// TIA Portal project "Vent_Fan_PLC_202203231" (V16)

(* hardware
DEVICE "ET 200SP station_1"  ET 200SP-Station
   slot 0: "Rack_0"  Rack  6ES5 710-8MAx1
   slot 1: "Roof Fans PLC"  CPU 1512SP-1 PN  6ES7 512-1DK01-0AB0  V2.1
      slot 32768: "PROFINET interface_1"  X1
         slot 32771: "Port_3"  X1 P3
   slot 2: "DI 16x24VDC ST_1"  DI 16x24VDC ST  6ES7 131-6BH00-0BA0  V1.1
      slot 1: "DI 16x24VDC ST_1"  DI 16x24VDC ST
   slot 3: "DQ 16x24VDC/0.5A ST_1"  DQ 16x24VDC/0.5A ST  6ES7 132-6BH00-0BA0  V1.0
      slot 1: "DQ 16x24VDC/0.5A ST_1"  DQ 16x24VDC/0.5A ST
   slot 4: "Server module_1"  Server module  6ES7 193-6PA00-0AA0  V1.1
      slot 1: "Server module_1"  Server module
   slot 127: "BA 2xRJ45"  BA 2xRJ45  6ES7 193-6AR00-0AA0  V0.0
      slot 32769: "Port_1"  X1 P1  6ES7 193-6AR00-0AA0
      slot 32770: "Port_2"  X1 P2  6ES7 193-6AR00-0AA0
DEVICE "SINAMICS G_1"  Sinamics.Device
   slot 0: "	_0"  Rail  SinamicsG120CRackP
   slot 0: "RTU-0035"  G120C PN  6SL3210-1KE15-8UF2  4.7.10
      slot 1: "PROFINET interface"  MDD-SinamicsG120-P
      slot 3: "PM G120C"  PM G120C  6SL3210-1KE15-8UF2  -
DEVICE "SINAMICS G_2"  Sinamics.Device
   slot 0: "	_0"  Rail  SinamicsG120CRackP
   slot 0: "RTU-0010"  G120C PN  6SL3210-1KE15-8UF2  4.7.10
      slot 1: "PROFINET interface"  MDD-SinamicsG120-P
      slot 3: "PM G120C"  PM G120C  6SL3210-1KE15-8UF2  -
DEVICE "SINAMICS G_3"  Sinamics.Device
   slot 0: "	_0"  Rail  SinamicsG120CRackP
   slot 0: "RTU-0011"  G120C PN  6SL3210-1KE15-8UF2  4.7.10
      slot 1: "PROFINET interface"  MDD-SinamicsG120-P
      slot 3: "PM G120C"  PM G120C  6SL3210-1KE15-8UF2  -
DEVICE "SINAMICS G_4"  Sinamics.Device
   slot 0: "	_0"  Rail  SinamicsG120CRackP
   slot 0: "RTU-0014"  G120C PN  6SL3210-1KE15-8UF2  4.7.10
      slot 1: "PROFINET interface"  MDD-SinamicsG120-P
      slot 3: "PM G120C"  PM G120C  6SL3210-1KE15-8UF2  -
DEVICE "SINAMICS G_5"  Sinamics.Device
   slot 0: "	_0"  Rail  SinamicsG120CRackP
   slot 0: "RTU-0015"  G120C PN  6SL3210-1KE15-8UF2  4.7.10
      slot 1: "PROFINET interface"  MDD-SinamicsG120-P
      slot 3: "PM G120C"  PM G120C  6SL3210-1KE15-8UF2  -
DEVICE "SINAMICS G_6"  Sinamics.Device
   slot 0: "	_0"  Rail  SinamicsG120CRackP
   slot 0: "RTU-0020"  G120C PN  6SL3210-1KE15-8UF2  4.7.10
      slot 1: "PROFINET interface"  MDD-SinamicsG120-P
      slot 3: "PM G120C"  PM G120C  6SL3210-1KE15-8UF2  -
DEVICE "SINAMICS G_7"  Sinamics.Device
   slot 0: "	_0"  Rail  SinamicsG120CRackP
   slot 0: "RTU-0021"  G120C PN  6SL3210-1KE15-8UF2  4.7.10
      slot 1: "PROFINET interface"  MDD-SinamicsG120-P
      slot 3: "PM G120C"  PM G120C  6SL3210-1KE15-8UF2  -
DEVICE "SINAMICS G_8"  Sinamics.Device
   slot 0: "	_0"  Rail  SinamicsG120CRackP
   slot 0: "RTU-0052"  G120C PN  6SL3210-1KE15-8UF2  4.7.10
      slot 1: "PROFINET interface"  MDD-SinamicsG120-P
      slot 3: "PM G120C"  PM G120C  6SL3210-1KE15-8UF2  -
DEVICE "SINAMICS G_9"  Sinamics.Device
   slot 0: "	_0"  Rail  SinamicsG120CRackP
   slot 0: "RTU-0053"  G120C PN  6SL3210-1KE15-8UF2  4.7.10
      slot 1: "PROFINET interface"  MDD-SinamicsG120-P
      slot 3: "PM G120C"  PM G120C  6SL3210-1KE15-8UF2  -
DEVICE "SINAMICS G_10"  Sinamics.Device
   slot 0: "	_0"  Rail  SinamicsG120CRackP
   slot 0: "RTU-0054"  G120C PN  6SL3210-1KE15-8UF2  4.7.10
      slot 1: "PROFINET interface"  MDD-SinamicsG120-P
      slot 3: "PM G120C"  PM G120C  6SL3210-1KE15-8UF2  -
DEVICE "SINAMICS G_11"  Sinamics.Device
   slot 0: "	_0"  Rail  SinamicsG120CRackP
   slot 0: "RTU-0055"  G120C PN  6SL3210-1KE15-8UF2  4.7.10
      slot 1: "PROFINET interface"  MDD-SinamicsG120-P
      slot 3: "PM G120C"  PM G120C  6SL3210-1KE15-8UF2  -
DEVICE "SINAMICS G_12"  Sinamics.Device
   slot 0: "	_0"  Rail  SinamicsG120CRackP
   slot 0: "RTU-0042"  G120C PN  6SL3210-1KE15-8UF2  4.7.10
      slot 1: "PROFINET interface"  MDD-SinamicsG120-P
      slot 3: "PM G120C"  PM G120C  6SL3210-1KE15-8UF2  -
*)

// ===== PLC "Roof Fans PLC"  CPU 1512SP-1 PN =====

VAR_GLOBAL   // PLC tag table "Default tag table"
   "System_Byte" AT %MB1 : Byte;
   "FirstScan" AT %M1.0 : Bool;
   "DiagStatusUpdate" AT %M1.1 : Bool;
   "AlwaysTRUE" AT %M1.2 : Bool;
   "AlwaysFALSE" AT %M1.3 : Bool;
   "Clock_Byte" AT %MB0 : Byte;
   "Clock_10Hz" AT %M0.0 : Bool;
   "Clock_5Hz" AT %M0.1 : Bool;
   "Clock_2.5Hz" AT %M0.2 : Bool;
   "Clock_2Hz" AT %M0.3 : Bool;
   "Clock_1.25Hz" AT %M0.4 : Bool;
   "Clock_1Hz" AT %M0.5 : Bool;
   "Clock_0.625Hz" AT %M0.6 : Bool;
   "Clock_0.5Hz" AT %M0.7 : Bool;
   "Drive_Temp" AT %MD100 : Real;
END_VAR

VAR_GLOBAL CONSTANT   // PLC tag table "Default tag table"
   "STATION_COUNT" : Int := 49;   // 0 indexed
   "SCHEDULES_PER_DAY" : Int := 4;   // 0 indexed
   "TIME_STRING_LENGTH" : Int := 20;   // standard indexed
END_VAR

VAR_GLOBAL   // PLC tag table "INPUTS"
   "Input_1" AT %I0.0 : Bool;
   "Input_2" AT %I0.2 : Bool;
   "Input_3" AT %I0.3 : Bool;
   "Input_4" AT %I0.4 : Bool;
   "Input_5" AT %I0.5 : Bool;
   "Input_6" AT %I0.6 : Bool;
   "Input_7" AT %I0.7 : Bool;
   "Input_8" AT %I1.0 : Bool;
   "Input_9" AT %I1.1 : Bool;
   "Input_10" AT %I1.2 : Bool;
   "Input_11" AT %I1.3 : Bool;
   "Input_12" AT %I1.4 : Bool;
   "Input_13" AT %I1.5 : Bool;
   "Input_14" AT %I1.6 : Bool;
   "Input_15" AT %I1.7 : Bool;
END_VAR

VAR_GLOBAL   // PLC tag table "OUTPUTS"
   "Output_1" AT %Q0.0 : Bool;
   "Output_15" AT %Q1.6 : Bool;
   "Output_2" AT %Q0.1 : Bool;
   "Output_3" AT %Q0.2 : Bool;
   "Output_4" AT %Q0.3 : Bool;
   "Output_5" AT %Q0.4 : Bool;
   "Output_6" AT %Q0.5 : Bool;
   "Output_7" AT %Q0.6 : Bool;
   "Output_8" AT %Q0.7 : Bool;
   "Output_9" AT %Q1.0 : Bool;
   "Output_10" AT %Q1.1 : Bool;
   "Output_11" AT %Q1.2 : Bool;
   "Output_12" AT %Q1.3 : Bool;
   "Output_13" AT %Q1.4 : Bool;
   "Output_14" AT %Q1.5 : Bool;
END_VAR

VAR_GLOBAL   // PLC tag table "RTU-0035"
   "RTU-0035_Temperature" AT %IW260 : Word;
   "RTU-0035_Speed" AT %IW258 : Word;
   "RTU-0035_Current" AT %IW262 : Word;
END_VAR

VAR_GLOBAL   // PLC tag table "RTU-0010"
   "RTU-0010_Temperature" AT %IW268 : Word;
   "RTU-0010_Speed" AT %IW266 : Word;
   "RTU-0010_Current" AT %IW270 : Word;
END_VAR

VAR_GLOBAL   // PLC tag table "RTU-0011"
   "RTU-0011_Temperature" AT %IW276 : Word;
   "RTU-0011_Speed" AT %IW274 : Word;
   "RTU-0011_Current" AT %IW278 : Word;
END_VAR

VAR_GLOBAL   // PLC tag table "RTU-0014"
   "RTU-0014_Temperature" AT %IW284 : Word;
   "RTU-0014_Speed" AT %IW282 : Word;
   "RTU-0014_Current" AT %IW286 : Word;
END_VAR

VAR_GLOBAL   // PLC tag table "RTU-0015"
   "RTU-0015_Temperature" AT %IW292 : Word;
   "RTU-0015_Speed" AT %IW290 : Word;
   "RTU-0015_Current" AT %IW294 : Word;
END_VAR

VAR_GLOBAL   // PLC tag table "RTU-0020"
   "RTU-0020_Temperature" AT %IW300 : Word;
   "RTU-0020_Speed" AT %IW298 : Word;
   "RTU-0020_Current" AT %IW302 : Word;
END_VAR

VAR_GLOBAL   // PLC tag table "RTU-0021"
   "RTU-0021_Temperature" AT %IW308 : Word;
   "RTU-0021_Speed" AT %IW2306 : Word;
   "RTU-0021_Current" AT %IW310 : Word;
END_VAR

VAR_GLOBAL   // PLC tag table "RTU-0052"
   "RTU-0052_Temperature" AT %IW316 : Word;
   "RTU-0052_Speed" AT %IW314 : Word;
   "RTU-0052_Current" AT %IW318 : Word;
END_VAR

VAR_GLOBAL   // PLC tag table "RTU-0053"
   "RTU-0053_Temperature" AT %IW324 : Word;
   "RTU-0053_Speed" AT %IW322 : Word;
   "RTU-0053_Current" AT %IW326 : Word;
END_VAR

VAR_GLOBAL   // PLC tag table "RTU-0054"
   "RTU-0054_Temperature" AT %IW332 : Word;
   "RTU-0054_Speed" AT %IW330 : Word;
   "RTU-0054_Current" AT %IW334 : Word;
END_VAR

VAR_GLOBAL   // PLC tag table "RTU-0055"
   "RTU-0055_Temperature" AT %IW340 : Word;
   "RTU-0055_Speed" AT %IW338 : Word;
   "RTU-0055_Current" AT %IW342 : Word;
END_VAR

VAR_GLOBAL   // PLC tag table "RTU-0042"
   "RTU-0042_Temperature" AT %IW348 : Word;
   "RTU-0042_Speed" AT %IW346 : Word;
   "RTU-0042_Current" AT %IW350 : Word;
END_VAR

TYPE "Web_Meta.UDT"
   STRUCT
      drive : "Drive.UDT";
      faults : "Faults.UDT";
      id : Int;
      manual : "Station.Web_Interface.Manual.UDT";
      selected_station : Int;
      scheduled_speed : Real;
      temporal_schedule : "Web_Meta.Web_Interface.Schedules.Temporal.UDT";
      thermal_schedule : "Schedules.Thermal.UDT";
   END_STRUCT;
END_TYPE

TYPE "Sensors.Thermal.UDT"
   STRUCT
      me : "Convert.Word_to_Real.UDT";
   END_STRUCT;
END_TYPE

TYPE "Sensors.UDT"
   STRUCT
      thermal : "Sensors.Thermal.UDT";
   END_STRUCT;
END_TYPE

TYPE "Drive.UDT"
   STRUCT
      commands : "Drive.Commands.UDT";
      commands_manual : "Drive.Commands.UDT";
      commands_thermal : "Drive.Commands.UDT";
      commands_temporal : "Drive.Commands.UDT";
      feedback : "Drive.Feedback.UDT";
      sensors : "Sensors.UDT";
   END_STRUCT;
END_TYPE

TYPE "Stations.UDT"
   STRUCT
      me : Array[0.."STATION_COUNT"] of "Station.UDT";
   END_STRUCT;
   // me[7].drive.sensors.thermal.me.processed := 76.8;
   // me[7].drive.feedback.speed.me.processed := 1100.56;
   // me[7].drive.feedback.current.me.processed := 3.78;
END_TYPE

TYPE "Station.UDT"
   STRUCT
      drive : "Drive.UDT";
      faults : "Faults.UDT";
      interface : "Interface.UDT";
      schedules : "Schedules.UDT";
   END_STRUCT;
END_TYPE

TYPE "Drive.Feedback.UDT"
   STRUCT
      faults : String := 'none';
      current : "Drive.Feedback.Current.UDT";
      speed : "Drive.Feedback.Speed.UDT";
      state : String := 'not running';
   END_STRUCT;
END_TYPE

TYPE "Convert.Word_to_Real.UDT"
   STRUCT
      raw : Word;
      processed : Real;
   END_STRUCT;
END_TYPE

TYPE "Drive.Feedback.Speed.UDT"
   STRUCT
      me : "Convert.Word_to_Real.UDT";
   END_STRUCT;
END_TYPE

TYPE "Drive.Feedback.Current.UDT"
   STRUCT
      me : "Convert.Word_to_Real.UDT";
   END_STRUCT;
END_TYPE

TYPE "Station.Web_Interface.UDT"
   STRUCT
      manual : "Station.Web_Interface.Manual.UDT";
      temporal : "Web_Meta.Web_Interface.Schedules.Temporal.UDT";
   END_STRUCT;
END_TYPE

TYPE "Station.Web_Interface.Manual.UDT"
   STRUCT
      acknowledge : Bool;
      command_speed : Real;
      mode : String[20] := 'stop';
      override : Bool;
      submit : Bool;
      toggle : Bool;
   END_STRUCT;
END_TYPE

TYPE "Schedules.Thermal.Element.UDT"
   STRUCT
      temperature : Real;
      speed : Real;
   END_STRUCT;
END_TYPE

TYPE "Schedules.Thermal.UDT"
   STRUCT
      start : "Schedules.Thermal.Element.UDT";
      max : "Schedules.Thermal.Element.UDT";
   END_STRUCT;
END_TYPE

TYPE "Schedules.UDT"
   STRUCT
      thermal : "Schedules.Thermal.UDT";
      temporal : "Schedules.Temporal.UDT";
   END_STRUCT;
END_TYPE

TYPE "Web_Meta.Web_Interface.Schedules.Temporal.Element.UDT"
   STRUCT
      start : String["TIME_STRING_LENGTH"];
      stop : String["TIME_STRING_LENGTH"];
      speed : Real;
   END_STRUCT;
END_TYPE

TYPE "Faults.UDT"
   STRUCT
      color : String[6];
      fault : String;
   END_STRUCT;
END_TYPE

TYPE "Interface.UDT"
   STRUCT
      current_feedback_b0 : DInt;
      id : USInt;
      raw_temp_sensor_b0 : DInt;
      sensor_max_temp : Real := 150.0;
      sensor_min_temp : Real;
      speed_feedback_b0 : DInt;
      max_speed : Real := 1500.0;
      profinet_pointer_to_drive : Hw_SubModule;
   END_STRUCT;
END_TYPE

TYPE "Interface.Thermal.UDT"
   STRUCT
      pointer_to_raw_value : DInt;   // input word number of data from drive
      min : Real;
      max : Real := 150.0;
   END_STRUCT;
END_TYPE

TYPE "Interface.Drive.Feedback.UDT"
   STRUCT
      current : DInt;   // pointer to input word with raw value
      speed : DInt;   // pointer to input word with raw value
   END_STRUCT;
END_TYPE

TYPE "Interface.Sensors.UDT"
   STRUCT
      thermal : "Interface.Thermal.UDT";
   END_STRUCT;
END_TYPE

TYPE "Drive.Commands.UDT"
   STRUCT
      override : Bool;
      run : Bool;
      speed : Real;
      stop : Bool;
   END_STRUCT;
END_TYPE

TYPE "Interface.Drive.Settings.UTD"
   STRUCT
      id : Bool;
      profinet_pointer_to_drive : Hw_SubModule;
      max_speed : Real := 1500.0;
   END_STRUCT;
END_TYPE

TYPE "OPC.Station.UDT"
   STRUCT
      current : Real;
      id : USInt;
      speed : Real;
      temperature : Real;
   END_STRUCT;
END_TYPE

TYPE "OPC.Stations.UDT"
   STRUCT
      me : Array[0.."STATION_COUNT"] of "OPC.Station.UDT";
   END_STRUCT;
END_TYPE

TYPE "Web_Meta.Web_Interface.Schedules.Temporal.UDT"
   STRUCT
      monday : Array[0.."SCHEDULES_PER_DAY"] of "Web_Meta.Web_Interface.Schedules.Temporal.Element.UDT";
      tuesday : Array[0.."SCHEDULES_PER_DAY"] of "Web_Meta.Web_Interface.Schedules.Temporal.Element.UDT";
      wednesday : Array[0.."SCHEDULES_PER_DAY"] of "Web_Meta.Web_Interface.Schedules.Temporal.Element.UDT";
      thursday : Array[0.."SCHEDULES_PER_DAY"] of "Web_Meta.Web_Interface.Schedules.Temporal.Element.UDT";
      friday : Array[0.."SCHEDULES_PER_DAY"] of "Web_Meta.Web_Interface.Schedules.Temporal.Element.UDT";
      saturday : Array[0.."SCHEDULES_PER_DAY"] of "Web_Meta.Web_Interface.Schedules.Temporal.Element.UDT";
      sunday : Array[0.."SCHEDULES_PER_DAY"] of "Web_Meta.Web_Interface.Schedules.Temporal.Element.UDT";
      new_data : Bool;
   END_STRUCT;
END_TYPE

TYPE "Schedules.Temporal.UDT"
   STRUCT
      monday : Array[0.."SCHEDULES_PER_DAY"] of "Schedules.Temporal.Element.UDT";
      tuesday : Array[0.."SCHEDULES_PER_DAY"] of "Schedules.Temporal.Element.UDT";
      wednesday : Array[0.."SCHEDULES_PER_DAY"] of "Schedules.Temporal.Element.UDT";
      thursday : Array[0.."SCHEDULES_PER_DAY"] of "Schedules.Temporal.Element.UDT";
      friday : Array[0.."SCHEDULES_PER_DAY"] of "Schedules.Temporal.Element.UDT";
      saturday : Array[0.."SCHEDULES_PER_DAY"] of "Schedules.Temporal.Element.UDT";
      sunday : Array[0.."SCHEDULES_PER_DAY"] of "Schedules.Temporal.Element.UDT";
   END_STRUCT;
END_TYPE

TYPE "Schedules.Temporal.Element.Date_Time.UDT"
   STRUCT
      month : USInt;
      day : USInt;
      weekday : USInt;
      hour : USInt;
      minute : USInt;
   END_STRUCT;
END_TYPE

TYPE "Schedules.Temporal.Element.UDT"
   STRUCT
      start : "Schedules.Temporal.Element.Date_Time.UDT";
      stop : "Schedules.Temporal.Element.Date_Time.UDT";
      speed : Real;
   END_STRUCT;
END_TYPE

DATA_BLOCK "Web_Meta"   // DB1
{ S7_Optimized_Access := 'TRUE' }
VERSION : 0.1
BEGIN
END_DATA_BLOCK

DATA_BLOCK "Stations"   // DB2
{ S7_Optimized_Access := 'TRUE' }
VERSION : 0.1
BEGIN
   me[7].interface.id := 42;
   me[0].interface.id := 10;
   me[1].interface.id := 11;
   me[2].interface.id := 14;
   me[8].interface.id := 52;
   me[3].interface.id := 15;
   me[5].interface.id := 21;
   me[6].interface.id := 35;
   me[4].interface.id := 20;
   me[9].interface.id := 53;
   me[10].interface.id := 54;
   me[11].interface.id := 55;
   me[6].interface.current_feedback_b0 := 262;
   me[6].interface.raw_temp_sensor_b0 := 260;
   me[6].interface.sensor_max_temp := 150.0;
   me[6].interface.speed_feedback_b0 := 258;
   me[6].interface.max_speed := 1500.0;
   me[6].interface.profinet_pointer_to_drive := 269;
   me[0].interface.current_feedback_b0 := 270;
   me[0].interface.raw_temp_sensor_b0 := 268;
   me[0].interface.speed_feedback_b0 := 266;
   me[0].interface.profinet_pointer_to_drive := 278;
   me[1].interface.profinet_pointer_to_drive := 287;
   me[1].interface.speed_feedback_b0 := 274;
   me[1].interface.raw_temp_sensor_b0 := 276;
   me[1].interface.current_feedback_b0 := 278;
   me[2].interface.speed_feedback_b0 := 282;
   me[2].interface.raw_temp_sensor_b0 := 284;
   me[2].interface.current_feedback_b0 := 286;
   me[2].interface.profinet_pointer_to_drive := 296;
   me[3].interface.profinet_pointer_to_drive := 305;
   me[4].interface.profinet_pointer_to_drive := 314;
   me[5].interface.profinet_pointer_to_drive := 323;
   me[10].interface.profinet_pointer_to_drive := 350;
   me[8].interface.profinet_pointer_to_drive := 332;
   me[9].interface.profinet_pointer_to_drive := 341;
   me[11].interface.profinet_pointer_to_drive := 359;
   me[3].interface.speed_feedback_b0 := 290;
   me[4].interface.speed_feedback_b0 := 298;
   me[5].interface.speed_feedback_b0 := 306;
   me[8].interface.speed_feedback_b0 := 314;
   me[9].interface.speed_feedback_b0 := 322;
   me[10].interface.speed_feedback_b0 := 330;
   me[11].interface.speed_feedback_b0 := 338;
   me[3].interface.raw_temp_sensor_b0 := 292;
   me[3].interface.current_feedback_b0 := 294;
   me[4].interface.raw_temp_sensor_b0 := 300;
   me[4].interface.current_feedback_b0 := 302;
   me[5].interface.raw_temp_sensor_b0 := 308;
   me[5].interface.current_feedback_b0 := 310;
   me[8].interface.raw_temp_sensor_b0 := 316;
   me[8].interface.current_feedback_b0 := 318;
   me[9].interface.raw_temp_sensor_b0 := 324;
   me[9].interface.current_feedback_b0 := 326;
   me[10].interface.raw_temp_sensor_b0 := 332;
   me[10].interface.current_feedback_b0 := 334;
   me[11].interface.raw_temp_sensor_b0 := 340;
   me[11].interface.current_feedback_b0 := 342;
   me[7].interface.raw_temp_sensor_b0 := 348;
   me[7].interface.current_feedback_b0 := 350;
   me[7].interface.speed_feedback_b0 := 346;
   me[7].interface.profinet_pointer_to_drive := 368;
END_DATA_BLOCK

DATA_BLOCK "All_Stations_IDB"   // DB3
{ S7_Optimized_Access := 'TRUE' }
VERSION : 0.1
// stored: InstanceOfName All_Stations
"All_Stations"
BEGIN
END_DATA_BLOCK

DATA_BLOCK "OPC.Stations"   // DB4
{ S7_Optimized_Access := 'TRUE' }
VERSION : 0.1
BEGIN
END_DATA_BLOCK

DATA_BLOCK "OPC_Map_IDB"   // DB5
{ S7_Optimized_Access := 'TRUE' }
VERSION : 0.1
// stored: InstanceOfName OPC_Map
"OPC_Map"
BEGIN
END_DATA_BLOCK

FUNCTION_BLOCK "Single_Station"   // FB1, SCL
{ S7_Optimized_Access := 'TRUE' }
VERSION : 0.1
   VAR_INPUT
      current_station : Int;
      selected_station : Int;
   END_VAR
   VAR_IN_OUT
      manual : "Station.Web_Interface.Manual.UDT";
      station : "Station.UDT";
   END_VAR
   VAR
      SinaSpeed : SinaSpeed;
   END_VAR
   VAR_TEMP
      _AxisEnabled : Bool;
      _DiagId : Word;
      _Lockout : Bool;
      _ActVelocity : Real;
      _Error : Bool;
      _Status : Word;
   END_VAR
BEGIN
   REGION "DRIVE"

       REGION "COMMANDS"
           "Drive.Commands"(current_station := #current_station,
                            selected_station := #selected_station,
                            thermal_sensor := #station.drive.sensors.thermal,
                            commands := #station.drive.commands,
                            commands_manual := #station.drive.commands_manual,
                            commands_temporal := #station.drive.commands_temporal,
                            commands_thermal := #station.drive.commands_thermal,
                            manual := #manual,
                            thermal := #station.schedules.thermal,
                            temporal := #station.schedules.temporal);
       END_REGION

       REGION "SEND COMMANDS"
           #SinaSpeed(EnableAxis := #station.drive.commands.run AND NOT #station.drive.commands.stop,
                      AckError := #manual.acknowledge,
                      SpeedSp := "Drive.Feedback.Speed.Percent_to_RPM"(as_percent := #station.drive.commands.speed, max_speed := #station.interface.max_speed),
                      RefSpeed := #station.interface.max_speed,
                      ConfigAxis := 16#3F,
                      HWIDSTW := #station.interface.profinet_pointer_to_drive,
                      HWIDZSW := #station.interface.profinet_pointer_to_drive,
                      AxisEnabled => #_AxisEnabled,
                      Lockout => #_Lockout,
                      ActVelocity => #_ActVelocity,
                      Error => #_Error,
                      Status => #_Status,
                      DiagId => #_DiagId);
           #manual.acknowledge := FALSE;
       END_REGION

       REGION "FEEDBACK"
           "Drive.Feedback"(pointer_to_current_feedback := #station.interface.current_feedback_b0,
                            pointer_to_speed_feedback := #station.interface.speed_feedback_b0,
                            feedback_data := #station.drive.feedback);
       END_REGION

       REGION "SENSORS"
           "Drive.Sensors"(pointer_to_raw_value := #station.interface.raw_temp_sensor_b0,
                           minimum_temperature := #station.interface.sensor_min_temp,
                           maximum_temperature := #station.interface.sensor_max_temp,
                           sensors := #station.drive.sensors);
       END_REGION

       REGION "FAULTS"
           "Faults"(fault_code := #_DiagId,
                    station := #station);
       END_REGION

   END_REGION
END_FUNCTION_BLOCK

FUNCTION_BLOCK "All_Stations"   // FB2, SCL
{ S7_Optimized_Access := 'TRUE' }
VERSION : 0.1
   VAR_IN_OUT
      stations : "Stations.UDT";
      web_meta : "Web_Meta.UDT";
   END_VAR
   VAR
      single_station : Array[0.."STATION_COUNT"] of "Single_Station";
      "Web_Meta.Load_Data" : "Web_Meta.Load_Data";
   END_VAR
   VAR_TEMP
      i : Int;
   END_VAR
BEGIN
   REGION "UPDATE WEB_META"
       IF #web_meta.selected_station <> -1 THEN
           #"Web_Meta.Load_Data"(selected_station := #web_meta.selected_station,
                                 id := #web_meta.id,
                                 faults := #web_meta.faults,
                                 drive := #web_meta.drive,
                                 manual := #web_meta.manual,
                                 stations := #stations,
                                 thermal_schedule := #web_meta.thermal_schedule,
                                 temporal_schedule := #web_meta.temporal_schedule);
       END_IF;

   END_REGION

   REGION "STATION DRIVERS"
       FOR #i := 0 TO "STATION_COUNT" DO
           IF #stations.me[#i].interface.id = 0 THEN
               CONTINUE;
           END_IF;
           #single_station[#i](current_station := #i,
                               selected_station := #web_meta.selected_station,
                               manual := #web_meta.manual,
                               station := #stations.me[#i]);
       END_FOR;
   END_REGION
END_FUNCTION_BLOCK

FUNCTION_BLOCK "Web_Meta.Load_Data"   // FB3, SCL
{ S7_Optimized_Access := 'TRUE' }
VERSION : 0.1
   VAR_INPUT
      selected_station : Int;
   END_VAR
   VAR_IN_OUT
      id : Int;
      faults : "Faults.UDT";
      drive : "Drive.UDT";
      manual : "Station.Web_Interface.Manual.UDT";
      stations : "Stations.UDT";
      thermal_schedule : "Schedules.Thermal.UDT";
      temporal_schedule : "Web_Meta.Web_Interface.Schedules.Temporal.UDT";
   END_VAR
   VAR
      _last_selected_station : Int;
   END_VAR
BEGIN
   #id := #stations.me[#selected_station].interface.id;
   #faults := #stations.me[#selected_station].faults;
   #thermal_schedule := #stations.me[#selected_station].schedules.thermal;
   #drive := #stations.me[#selected_station].drive;
   IF #_last_selected_station = #selected_station THEN
       "Web_Meta.Update_Temporal.Web_to_PLC"(web := #temporal_schedule,
                                             plc := #stations.me[#selected_station].schedules.temporal);
   END_IF;
   IF #_last_selected_station <> #selected_station THEN
       "Web_Meta.Update_Manual.PLC_to_Web"(station := #stations.me[#selected_station],
                                           manual := #manual);
       "Web_Meta.Update_Temporal.PLC_to_Web"(plc := #stations.me[#selected_station].schedules.temporal,
                                             web := #temporal_schedule);
   END_IF;
   #_last_selected_station := #selected_station;
END_FUNCTION_BLOCK

FUNCTION_BLOCK "OPC_Map"   // FB4, SCL
{ S7_Optimized_Access := 'TRUE' }
VERSION : 0.1
   VAR_INPUT
      stations : "Stations.UDT";
   END_VAR
   VAR_IN_OUT
      "opc.stations" : "OPC.Stations.UDT";
   END_VAR
   VAR_TEMP
      _length : Int;
      _i : Int;
   END_VAR
BEGIN
   #_length := UDINT_TO_INT("Array.Any.Length"(#stations.me));
   FOR #_i := 0 TO #_length - 1 DO
       "OPC_Map.Map_Station"(station:=#stations.me[#_i],
                             "opc.station":=#"opc.stations".me[#_i]);
   END_FOR;
END_FUNCTION_BLOCK

FUNCTION "Word.ToString" : String   // FC1, SCL
{ S7_Optimized_Access := 'TRUE' }
VERSION : 0.1
   VAR_INPUT
      value : Word;
   END_VAR
   VAR_TEMP
      _ret : String;
   END_VAR
BEGIN
   #"Word.ToString" := CONCAT_STRING(IN1 := "Byte.ToString"(#value.%B1),
                                     IN2 := "Byte.ToString"(#value.%B0));
END_FUNCTION

FUNCTION "Drive.Scale_Parameter" : Real   // FC2, SCL
{ S7_Optimized_Access := 'TRUE' }
VERSION : 0.1
   VAR_INPUT
      x_min : Word;
      x_max : Word;
      x_actual : Word;
      y_min : Real;
      y_max : Real;
   END_VAR
   VAR_TEMP
      x_real : Struct
         min : Real;
         max : Real;
         actual : Real;
      END_STRUCT;
   END_VAR
BEGIN
   #x_real.min := INT_TO_REAL(WORD_TO_INT(#x_min));
   #x_real.max := INT_TO_REAL(WORD_TO_INT(#x_max));
   #x_real.actual := INT_TO_REAL(WORD_TO_INT(#x_actual));
   #"Drive.Scale_Parameter" := (#y_max - #y_min) /  (#x_real.max - #x_real.min) * (#x_real.actual - #x_real.min)  + #y_min;
END_FUNCTION

FUNCTION "Drive.Feedback" : Void   // FC3, SCL
{ S7_Optimized_Access := 'TRUE' }
VERSION : 0.1
   VAR_INPUT
      pointer_to_current_feedback : DInt;
      pointer_to_speed_feedback : DInt;
   END_VAR
   VAR_IN_OUT
      feedback_data : "Drive.Feedback.UDT";
   END_VAR
BEGIN
   REGION "CURRENT"
       #feedback_data.current := "Drive.Feedback.Current"(#pointer_to_current_feedback);
   END_REGION

   REGION "SPEED"
       #feedback_data.speed := "Drive.Feedback.Speed"(pointer_to_raw := #pointer_to_speed_feedback);
   END_REGION

   REGION "STATE"
       #feedback_data.state := "Drive.Feedback.State"(#feedback_data.speed);
   END_REGION
END_FUNCTION

FUNCTION "Drive.Sensors" : Void   // FC4, SCL
{ S7_Optimized_Access := 'TRUE' }
VERSION : 0.1
   VAR_INPUT
      pointer_to_raw_value : DInt;
      minimum_temperature : Real;
      maximum_temperature : Real;
   END_VAR
   VAR_IN_OUT
      sensors : "Sensors.UDT";
   END_VAR
BEGIN
   REGION "TEMPERATURE"
       #sensors.thermal := "Drive.Sensors.Thermal"(pointer_to_raw_value := #pointer_to_raw_value,
                                                   minimum_temperature := #minimum_temperature,
                                                   maximum_temperature := #maximum_temperature);
   END_REGION
END_FUNCTION

FUNCTION "Drive.Feedback.Current" : "Drive.Feedback.Current.UDT"   // FC5, SCL
{ S7_Optimized_Access := 'TRUE' }
VERSION : 0.1
   VAR_INPUT
      pointer_to_current : DInt;
   END_VAR
   VAR_TEMP
      _ret : "Drive.Feedback.Current.UDT";
   END_VAR
   VAR CONSTANT
      INPUT_AREA : Byte := 16#81;
      AREA_NOT_A_DB : DInt;
      MAX_WORD : Word := 16#4000;
      MIN_WORD : Word;
      MAX_CURRENT : Real := 6.3;
      MIN_CURRENT : Real;
   END_VAR
BEGIN
   #_ret.me.raw := PEEK_WORD(area := #INPUT_AREA,
                             dbNumber := #AREA_NOT_A_DB,
                             byteOffset := #pointer_to_current);
   #_ret.me.processed := "Drive.Scale_Parameter"(x_min := #MAX_WORD,
                                                 x_max := #MIN_WORD,
                                                 x_actual := #_ret.me.raw,
                                                 y_min := #MAX_CURRENT,
                                                 y_max := #MIN_CURRENT);
   #"Drive.Feedback.Current" := #_ret;
END_FUNCTION

FUNCTION "Drive.Feedback.Speed" : "Drive.Feedback.Speed.UDT"   // FC6, SCL
{ S7_Optimized_Access := 'TRUE' }
VERSION : 0.1
   VAR_INPUT
      pointer_to_raw : DInt;
   END_VAR
   VAR_TEMP
      _ret : "Drive.Feedback.Speed.UDT";
   END_VAR
   VAR CONSTANT
      INPUT_AREA : Byte := 16#81;
      AREA_NOT_A_DB : DInt;
      MIN_SPEED : Word := 16#00_00;
      MAX_SPEED : Word := 16#40_00;
   END_VAR
BEGIN
   #_ret.me.raw := PEEK_WORD(area := #INPUT_AREA,
                             dbNumber := #AREA_NOT_A_DB,
                             byteOffset := #pointer_to_raw);
   #_ret.me.processed := "Drive.Scale_Parameter"(x_min := #MIN_SPEED,
                                                 x_max := #MAX_SPEED,
                                                 x_actual := #_ret.me.raw,
                                                 y_min := 0,
                                                 y_max := 100.0); 
   #"Drive.Feedback.Speed" := #_ret;
END_FUNCTION

FUNCTION "Drive.Sensors.Thermal" : "Sensors.Thermal.UDT"   // FC7, SCL
{ S7_Optimized_Access := 'TRUE' }
VERSION : 0.1
   VAR_INPUT
      pointer_to_raw_value : DInt;
      minimum_temperature : Real;
      maximum_temperature : Real;
   END_VAR
   VAR_TEMP
      _ret : "Sensors.Thermal.UDT";
   END_VAR
   VAR CONSTANT
      SENSOR_MAX : Word := 16#3F_FF;
      SENSOR_MIN : Word;
      INPUT_AREA : Byte := 16#81;
      AREA_NOT_A_DB : DInt;
   END_VAR
BEGIN
   #_ret.me.raw := PEEK_WORD(area := #INPUT_AREA,
                             dbNumber := #AREA_NOT_A_DB,
                             byteOffset := #pointer_to_raw_value);
   #_ret.me.processed := "Drive.Scale_Parameter"(x_min := #SENSOR_MIN,
                                                     x_max := #SENSOR_MAX,
                                                     x_actual := #_ret.me.raw,
                                                     y_min := #minimum_temperature,
                                                     y_max := #maximum_temperature);
   #"Drive.Sensors.Thermal" := #_ret;
END_FUNCTION

FUNCTION "Drive.Feedback.State" : String   // FC8, SCL
{ S7_Optimized_Access := 'TRUE' }
VERSION : 0.1
   VAR_INPUT
      speed : "Drive.Feedback.Speed.UDT";
   END_VAR
   VAR_TEMP
      _ret : String;
   END_VAR
   VAR CONSTANT
      NOT_RUNNING : String := 'not running';
      RUNNING : String := 'running';
   END_VAR
BEGIN
   IF #speed.me.processed = 0.0 THEN
       #"Drive.Feedback.State" := #NOT_RUNNING;
       RETURN;
   END_IF;
   #"Drive.Feedback.State" := #RUNNING;
END_FUNCTION

FUNCTION "Drive.Commands.Run.Thermal" : Void   // FC9, SCL
{ S7_Optimized_Access := 'TRUE' }
VERSION : 0.1
   VAR_INPUT
      sensor : "Sensors.Thermal.UDT";
      schedule : "Schedules.Thermal.UDT";
   END_VAR
   VAR_IN_OUT
      commands : "Drive.Commands.UDT";
   END_VAR
BEGIN
   REGION "TOO COLD"
       IF #sensor.me.processed < #schedule.start.temperature THEN
           #commands.run := FALSE;
           #commands.stop := TRUE;
           #commands.speed := 0.0;
           RETURN;
       END_IF;
   END_REGION


   REGION "TOO HOT"
       IF #sensor.me.processed > #schedule.max.temperature THEN
           #commands.run := TRUE;
           #commands.stop := FALSE;
           #commands.speed :=#schedule.max.speed;
           RETURN;
       END_IF;
   END_REGION


   REGION "JUST RIGHT"
       #commands.run := TRUE;
       #commands.stop := FALSE;
       #commands.speed := "Real.Scale"(x_min := #schedule.start.temperature,
                                       x_max := #schedule.max.temperature,
                                       x_actual := #sensor.me.processed,
                                       y_min := #schedule.start.speed,
                                       y_max := #schedule.max.speed);
   END_REGION
END_FUNCTION

FUNCTION "Drive.Commands.Run.Manual" : Void   // FC10, SCL
{ S7_Optimized_Access := 'TRUE' }
VERSION : 0.1
   VAR_IN_OUT
      web_manual : "Station.Web_Interface.Manual.UDT";
      commands : "Drive.Commands.UDT";
   END_VAR
   VAR CONSTANT
      _RUN : String := 'run';
      _STOP : String := 'stop';
      _OVERRIDE : String := 'override';
   END_VAR
BEGIN
   "Drive.Commands.Run.Manual.Override"(web_manual := #web_manual,
                                        commands := #commands);
   IF #web_manual.mode <> #_OVERRIDE THEN
       "Drive.Commands.Run.Manual.Mode"(web_manual := #web_manual,
                                        commands := #commands);
   END_IF;
END_FUNCTION

FUNCTION "Schedule.In_Schedule" : Real   // FC11, SCL
{ S7_Optimized_Access := 'TRUE' }